screen "1牵伸相关" 1280x740, template "模板_调试"
   on GenerateScreen: "TitleUpdater"()
   IOField "IO 域_5" at 461,39 size 126x56; FormatPattern 9.999
      ProcessValue <- "ST_Cam5_Data_Var_g_tz3"
   IOField "IO 域_10" at 181,306 size 114x56; FormatPattern 9.9999
      ProcessValue <- "ST_Cam5_Data_Var_fi"
   IOField "IO 域_11" at 181,235 size 126x55; FormatPattern s9.99
      ProcessValue <- "ST_Cam5_Data_Var_g_ratioV"
   IOField "IO 域_12" at 321,235 size 126x55; FormatPattern 9.99
      ProcessValue <- "ST_Cam5_Data_Var_g_ratioT"
   TextField "文本域_13" at 181,193 size 132x43; Text 'ratioV'
   TextField "文本域_14" at 321,193 size 132x43; Text 'ratioT'
   IOField "IO 域_14" at 461,235 size 126x55; FormatPattern 9.99
      ProcessValue <- "ST_Cam5_Data_Var_g_ratio"
   TextField "文本域_16" at 461,193 size 116x43; Text 'ratio'
   IOField "IO 域_7" at 181,39 size 126x56; FormatPattern 9999
      ProcessValue <- "ST_HMI_Var_HMI_r64Position_ChuChe"
   IOField "IO 域_9" at 181,123 size 126x56; FormatPattern 9.99
      ProcessValue <- "ST_HMI_Var_HMI_r64QianShen_All"
   IOField "IO 域_13" at 321,123 size 126x56; FormatPattern 9.99
      ProcessValue <- "ST_HMI_Var_HMI_r64QianShen_First"
   IOField "IO 域_15" at 461,123 size 126x56; FormatPattern 999
      ProcessValue <- "ST_HMI_Var_HMI_r64QianShen_FirstArea"
   IOField "IO 域_16" at 601,123 size 126x56; FormatPattern 99
      ProcessValue <- "ST_HMI_Var_HMI_r64QianShen_finalArea"
   Button "Button" at 615,39 size 98x56; TextOff 'CAM5'
      Appearance <- "Cam_5_accessState"
   IOField "IO 域_8" at 321,39 size 126x56; FormatPattern 999
      ProcessValue <- "ST_Cam5_Data_Var_g_vm"
   IOField "IO 域_1" at 968,39 size 126x56; FormatPattern 9999999999
      ProcessValue <- "ST_HMI_Var_HMI_i32_ZouChe_ZhanJu_ss_1"
   IOField "IO 域_2" at 968,111 size 126x56; FormatPattern 9999
      ProcessValue <- "ST_HMI_Var_HMI_r64_ZouChe_ZhanJu_Max_20"
      Visibility <- "ST_HMI_Var_HMI_bo_ZouChe_ZhanJu_Select"
   IOField "IO 域_3" at 968,183 size 126x56; FormatPattern 9999
      ProcessValue <- "ST_HMI_Var_HMI_r64_ZouChe_ZhanJu_Max_25"
      Visibility <- "ST_HMI_Var_HMI_bo_ZouChe_ZhanJu_Select"
   IOField "IO 域_4" at 968,255 size 126x56; FormatPattern 9999
      ProcessValue <- "ST_HMI_Var_HMI_r64_ZouChe_ZhanJu_Max_30"
      Visibility <- "ST_HMI_Var_HMI_bo_ZouChe_ZhanJu_Select"
   IOField "IO 域_6" at 968,327 size 126x56; FormatPattern 9999
      ProcessValue <- "ST_HMI_Var_HMI_r64_ZouChe_ZhanJu_Max_35"
      Visibility <- "ST_HMI_Var_HMI_bo_ZouChe_ZhanJu_Select"
   IOField "IO 域_17" at 968,399 size 126x56; FormatPattern 9999
      ProcessValue <- "ST_HMI_Var_HMI_r64_ZouChe_ZhanJu_Max_40"
      Visibility <- "ST_HMI_Var_HMI_bo_ZouChe_ZhanJu_Select"
   IOField "IO 域_18" at 968,471 size 126x56; FormatPattern 9999
      ProcessValue <- "ST_HMI_Var_HMI_r64_ZouChe_ZhanJu_Max_45"
      Visibility <- "ST_HMI_Var_HMI_bo_ZouChe_ZhanJu_Select"
   IOField "IO 域_19" at 968,543 size 126x56; FormatPattern 9999
      ProcessValue <- "ST_HMI_Var_HMI_r64_ZouChe_ZhanJu_Max_Effect"
      Visibility <- "ST_HMI_Var_HMI_bo_ZouChe_ZhanJu_Select"
   Button "Button_1" at 824,111 size 126x56; TextOff '2.0米'
      on Release: SetTag("ST_HMI_Var_HMI_i16_ZouChe_ZhanJu_Select", 20)
      Visibility <- "ST_HMI_Var_HMI_bo_ZouChe_ZhanJu_Select"
      Appearance <- "ST_HMI_Var_HMI_i16_ZouChe_ZhanJu_Select"
   Button "Button_2" at 824,183 size 126x56; TextOff '2.5米'
      on Release: SetTag("ST_HMI_Var_HMI_i16_ZouChe_ZhanJu_Select", 25)
      Visibility <- "ST_HMI_Var_HMI_bo_ZouChe_ZhanJu_Select"
      Appearance <- "ST_HMI_Var_HMI_i16_ZouChe_ZhanJu_Select"
   Button "Button_3" at 824,255 size 126x56; TextOff '3.0米'
      on Release: SetTag("ST_HMI_Var_HMI_i16_ZouChe_ZhanJu_Select", 30)
      Visibility <- "ST_HMI_Var_HMI_bo_ZouChe_ZhanJu_Select"
      Appearance <- "ST_HMI_Var_HMI_i16_ZouChe_ZhanJu_Select"
   Button "Button_4" at 824,327 size 126x56; TextOff '3.5米'
      on Release: SetTag("ST_HMI_Var_HMI_i16_ZouChe_ZhanJu_Select", 35)
      Visibility <- "ST_HMI_Var_HMI_bo_ZouChe_ZhanJu_Select"
      Appearance <- "ST_HMI_Var_HMI_i16_ZouChe_ZhanJu_Select"
   Button "Button_5" at 824,399 size 126x56; TextOff '4.0米'
      on Release: SetTag("ST_HMI_Var_HMI_i16_ZouChe_ZhanJu_Select", 40)
      Visibility <- "ST_HMI_Var_HMI_bo_ZouChe_ZhanJu_Select"
      Appearance <- "ST_HMI_Var_HMI_i16_ZouChe_ZhanJu_Select"
   Button "Button_6" at 824,471 size 126x56; TextOff '4.5米'
      on Release: SetTag("ST_HMI_Var_HMI_i16_ZouChe_ZhanJu_Select", 45)
      Visibility <- "ST_HMI_Var_HMI_bo_ZouChe_ZhanJu_Select"
      Appearance <- "ST_HMI_Var_HMI_i16_ZouChe_ZhanJu_Select"
   Button "Button_7" at 824,543 size 126x56; TextOff '生效'
      Visibility <- "ST_HMI_Var_HMI_bo_ZouChe_ZhanJu_Select"
   Button "Button_8" at 181,525 size 126x56; TextOff '2.0米'; TextList "Text_list_IP_Local_Remote_Select"
      on Release: InvertBit("ST_2_HMI_bo_IP_Local_remote_Select")
      Visibility <- "ST_HMI_Var_HMI_bo_ZouChe_ZhanJu_Select"
      Appearance <- "ST_2_HMI_bo_IP_Local_remote_Select"
      ProcessValue <- "ST_2_HMI_bo_IP_Local_remote_Select"
   IOField "IO 域_21" at 327,525 size 64x56; FormatPattern 999
      ProcessValue <- "ST_2_vIPArray{0}"
      Visibility <- "ST_HMI_Var_HMI_bo_ZouChe_ZhanJu_Select"
   IOField "IO 域_22" at 398,525 size 64x56; FormatPattern 999
      ProcessValue <- "ST_2_vIPArray{1}"
      Visibility <- "ST_HMI_Var_HMI_bo_ZouChe_ZhanJu_Select"
   IOField "IO 域_23" at 470,525 size 64x56; FormatPattern 999
      ProcessValue <- "ST_2_vIPArray{2}"
      Visibility <- "ST_HMI_Var_HMI_bo_ZouChe_ZhanJu_Select"
   IOField "IO 域_24" at 542,525 size 64x56; FormatPattern 999
      ProcessValue <- "ST_2_vIPArray{3}"
      Visibility <- "ST_HMI_Var_HMI_bo_ZouChe_ZhanJu_Select"
   Button "Button_9" at 181,432 size 126x56; TextOff '设备ID'; TextList "Text_list_IP_Local_Remote_Select"
      Appearance <- "ST_2_HMI_bo_IP_Local_remote_Select"
      Visibility <- "ST_HMI_Var_HMI_bo_ZouChe_ZhanJu_Select"
      ProcessValue <- "ST_2_HMI_bo_IP_Local_remote_Select"
   IOField "IO 域_20" at 328,432 size 135x56; FormatPattern 9999
      ProcessValue <- "ST_HMI_Var_HMI_u32_DeviceID"
      Visibility <- "ST_HMI_Var_HMI_bo_ZouChe_ZhanJu_Select"

screen "2加捻相关" 1280x740, template "模板_调试"
   on GenerateScreen: "TitleUpdater"()
   TextField "Text Field_58" at 327,45 size 304x42; Text '锭子加捻加速度'
   TextField "Text Field_1" at 168,8 size 156x23; Text '一、锭子加捻TO参数:'
   TextField "Text Field_60" at 327,101 size 304x42; Text '锭子加捻正起始加加速度'
   TextField "Text Field_61" at 327,157 size 304x42; Text '锭子加捻正终止加加速度'
   TextField "Text Field_62" at 327,213 size 304x42; Text '锭子加捻负起始加加速度'
   TextField "Text Field_63" at 327,269 size 304x42; Text '锭子加捻负终止加加速度'
   TextField "Text Field_66" at 327,325 size 304x42; Text '锭子点动加捻加速度'
   IOField "IO Field_38" at 194,41 size 112x42; FormatPattern 99999
      ProcessValue <- "ST_HMI_Var_HMI_r64Axis_DingZi_PositiveAccel_JiaNian"
   IOField "IO Field_40" at 194,97 size 112x42; FormatPattern 99999
      ProcessValue <- "ST_HMI_Var_HMI_r64Axis_DingZi_Positiveaccelstartjerk_JiaNian"
   IOField "IO Field_41" at 194,153 size 112x42; FormatPattern 99999
      ProcessValue <- "ST_HMI_Var_HMI_r64Axis_DingZi_positiveaccelendjerk_JiaNian"
   IOField "IO Field_42" at 194,209 size 112x42; FormatPattern 99999
      ProcessValue <- "ST_HMI_Var_HMI_r64Axis_DingZi_negativeaccelstartjerk_JiaNian"
   IOField "IO Field_43" at 194,265 size 112x42; FormatPattern 99999
      ProcessValue <- "ST_HMI_Var_HMI_r64Axis_DingZi_negativeaccelendjerk_JiaNian"
   IOField "IO Field_44" at 194,321 size 112x42; FormatPattern 99999
      ProcessValue <- "ST_HMI_Var_HMI_r64AccVelocity_Jog_JiaNian"

screen "3退绕相关1" 1280x740, template "模板_调试"
   on GenerateScreen: "TitleUpdater"()
   TextField "Text Field_58" at 153,27 size 668x41; Text '1.退绕成形弓速度————————————'
   TextField "Text Field_59" at 153,77 size 668x41; Text '2.退绕成形弓加速度————————————'
   TextField "Text Field_60" at 153,128 size 668x40; Text '3.退绕成形弓正向开始加加速度————————————'
   TextField "Text Field_61" at 153,178 size 668x41; Text '4.退绕成形弓正向结束加加速度————————————'
   TextField "Text Field_62" at 153,229 size 668x40; Text '5.退绕成形弓反向开始加加速度————————————'
   TextField "Text Field_1" at 153,5 size 247x26; Text '一、退绕成形弓TO参数:'
   TextField "Text Field_63" at 153,279 size 668x41; Text '6.退绕成形弓反向结束加加速度————————————'
   TextField "Text Field_41" at 153,361 size 668x41; Text '1.退绕结束纱线提前角度（越大，卷绕时，包络层螺距越大）—————————————————————'
   TextField "Text Field_42" at 153,413 size 668x41; Text '2.退绕开始位置—————————————————————————————'
   TextField "Text Field_43" at 153,465 size 668x41; Text '3.退绕结束位置—————————————————————————'
   TextField "Text Field_44" at 153,517 size 668x41; Text '4.退绕拐点比例———————————————————————————'
   TextField "Text Field_45" at 153,569 size 668x41; Text '5.退绕拐点点数---------------------'
   TextField "Text Field_3" at 153,327 size 260x26; Text '二、Cam_3曲线计算参数:'
   TextField "Text Field_46" at 153,621 size 668x41; Text '6.退绕圈数比例（越大，圈数越多，一般以0.03为单位调整）---------------------'
   IOField "IO Field_39" at 819,23 size 109x41; FormatPattern 9999
      ProcessValue <- "ST_HMI_Var_HMI_r64Axis_ChengXing_Velocity_TuiRao"
   IOField "IO Field_43" at 819,74 size 109x41; FormatPattern 9999
      ProcessValue <- "ST_HMI_Var_HMI_r64Axis_ChengXing_PositiveAccel_TuiRao"
   IOField "IO Field_44" at 819,125 size 109x41; FormatPattern 9999
      ProcessValue <- "ST_HMI_Var_HMI_r64Axis_ChengXing_positiveaccelstartjerk_TuiRao"
   IOField "IO Field_45" at 819,177 size 109x41; FormatPattern 9999
      ProcessValue <- "ST_HMI_Var_HMI_r64Axis_ChengXing_positiveaccelendjerk_TuiRao"
   IOField "IO Field_46" at 819,228 size 109x41; FormatPattern 9999
      ProcessValue <- "ST_HMI_Var_HMI_r64Axis_ChengXing_negativeaccelstartjerk_TuiRao"
   IOField "IO Field_47" at 819,280 size 109x40; FormatPattern 9999
      ProcessValue <- "ST_HMI_Var_HMI_r64Axis_ChengXing_negativeaccelendjerk_TuiRao"
   IOField "IO Field_53" at 819,367 size 109x41; FormatPattern 9999
      ProcessValue <- "ST_HMI_Var_HMI_alpha_TuiRao_5"
   IOField "IO Field_54" at 819,468 size 109x41; FormatPattern 99999
      ProcessValue <- "ST_HMI_Var_HMI_x_TuiRao_5"
   IOField "IO Field_55" at 819,570 size 109x41; FormatPattern 99
      ProcessValue <- "ST_HMI_Var_HMI_n_Change_TuiRao"
   IOField "IO Field_56" at 819,417 size 109x41; FormatPattern 9999
      ProcessValue <- "ST_HMI_Var_HMI_x_TuiRao_0"
   IOField "IO Field_57" at 819,519 size 109x41; FormatPattern 9.99
      ProcessValue <- "ST_HMI_Var_HMI_k_TuiRao"
   IOField "IO Field_58" at 819,621 size 109x41; FormatPattern 9.99
      ProcessValue <- "ST_HMI_Var_HMI_scalevalue_Cam_3"

screen "4退绕相关2" 1280x740, template "模板_调试"
   on GenerateScreen: "TitleUpdater"()
   TextField "Text Field_48" at 151,98 size 786x42; Text '2.退绕锭子响应正向加速度————————————————————'
   TextField "Text Field_49" at 151,154 size 786x42; Text '3.退绕锭子响应反向加速度————————————————————————'
   TextField "Text Field_1" at 151,9 size 204x27; Text '三、cam_3 TO参数'
   TextField "Text Field_65" at 151,42 size 786x42; Text '1.退绕锭子响应速度————————————————————'
   TextField "Text Field_4" at 151,210 size 235x27; Text '四、退绕张力TO参数'
   TextField "Text Field_54" at 151,309 size 786x42; Text '2.退绕张力加速度比例————————————————————'
   TextField "Text Field_66" at 151,253 size 786x42; Text '1.退绕张力速度比例————————————————————'
   TextField "Text Field_5" at 151,407 size 377x27; Text '五、退绕工艺进程衔接紧密性参数:'
   TextField "Text Field_63" at 151,449 size 786x42; Text '1.退绕锭子速度减少值————————————————————'
   TextField "Text Field_64" at 151,505 size 786x42; Text '2.开始退绕锭子速度————————————'
   IOField "IO Field_40" at 935,42 size 112x42; FormatPattern 9999
      ProcessValue <- "ST_HMI_Var_HMI_r64_cam_DingZi_velocity_TuiRao"
   IOField "IO Field_43" at 935,98 size 112x42; FormatPattern 99999
      ProcessValue <- "ST_HMI_Var_HMI_r64_cam_DingZi_positiveaccel_TuiRao"
   IOField "IO Field_47" at 935,154 size 112x42; FormatPattern 99999
      ProcessValue <- "ST_HMI_Var_HMI_r64_cam_DingZi_negativeaccel_TuiRao"
   IOField "IO Field_50" at 935,253 size 112x42; FormatPattern 9.99
      ProcessValue <- "ST_HMI_Var_HMI_r64Axis_1_ZhangLi_Velocity_from_ChengXing_ratio_tuirao"
   IOField "IO Field_51" at 935,309 size 112x42; FormatPattern 9.99
      ProcessValue <- "ST_HMI_Var_HMI_r64Axis_1_ZhangLi_PositiveAccel_from_ChengXing_ratio_tuirao"
   IOField "IO Field_52" at 935,449 size 112x42; FormatPattern 9999
      ProcessValue <- "ST_HMI_Var_HMI_r64Axis_DingZi_Velocity_JianShaoZhi"
   IOField "IO Field_53" at 935,505 size 112x42; FormatPattern 99
      ProcessValue <- "ST_HMI_Var_HMI_r64Axis_DingZi_Velocity_Start_TuiRao"
   IOField "IO Field_56" at 935,365 size 112x42; FormatPattern 9.99
      ProcessValue <- "ST_HMI_Var_HMI_r64Axis_1_ZhangLi_Additive_Torque_TuiRao"

screen "5成形相关" 1280x740, template "模板_调试"
   on GenerateScreen: "TitleUpdater"()
   TextField "Text Field_1" at 140,1 size 267x29; Text '一、成形凸轮曲线计算参数:'
   TextField "Text Field_58" at 138,36 size 648x39; Text '1.卷绕提前角度1——————————————————————'
   TextField "Text Field_59" at 138,81 size 648x40; Text '2.卷绕提前角度2——————————————————————————'
   TextField "Text Field_60" at 138,127 size 648x40; Text '3.卷绕提前角度3——————————————————————————'
   TextField "Text Field_61" at 138,174 size 648x40; Text '4.生头开始上锥体高度修正值——————————————————————————'
   TextField "Text Field_62" at 138,220 size 648x39; Text '5.最大直径时上椎体高度修正值——————————————————————————'
   TextField "Text Field_63" at 139,266 size 648x39; Text '6.满纱时上椎体高度修正值————————————————————————'
   TextField "Text Field_2" at 140,308 size 165x29; Text '二、cam1TO参数:'
   TextField "Text Field_64" at 140,337 size 648x39; Text '1.卷绕成形响应速度——————————————————————'
   TextField "Text Field_65" at 140,385 size 648x40; Text '2.卷绕成形响应正向加速度——————————————————————————'
   TextField "Text Field_66" at 140,435 size 648x40; Text '3.卷绕成形响应负向加速度——————————————————————————'
   TextField "Text Field_67" at 140,485 size 648x40; Text '4.卷绕成形响应正向开始加加速度——————————————————————————'
   TextField "Text Field_68" at 140,535 size 648x39; Text '5.卷绕成形响应正向结束加加速度——————————————————————————'
   TextField "Text Field_69" at 140,584 size 649x39; Text '6.卷绕成形响应反向开始加加速度————————————————————————'
   TextField "Text Field_70" at 140,633 size 648x40; Text '7.卷绕成形响应反向结束加加速度————————————————————————'
   IOField "IO Field_51" at 786,32 size 106x40; FormatPattern 99.9
      ProcessValue <- "ST_HMI_Var_HMI_alpha_JuanRao_1"
   IOField "IO Field_52" at 786,337 size 106x39; FormatPattern 9999
      ProcessValue <- "ST_HMI_Var_HMI_r64_cam_ChengXing_velocity_juanrao"
   IOField "IO Field_53" at 786,79 size 106x40; FormatPattern 99.9
      ProcessValue <- "ST_HMI_Var_HMI_alpha_JuanRao_2"
   IOField "IO Field_54" at 786,126 size 106x40; FormatPattern 99.9
      ProcessValue <- "ST_HMI_Var_HMI_alpha_JuanRao_3"
   IOField "IO Field_55" at 786,173 size 106x39; FormatPattern 99.9
      ProcessValue <- "ST_HMI_Var_HMI_r64_Hs2_0_delt"
   IOField "IO Field_56" at 786,219 size 106x39; FormatPattern 99.9
      ProcessValue <- "ST_HMI_Var_HMI_r64_Hs2_D_delt"
   IOField "IO Field_57" at 786,266 size 106x40; FormatPattern 99.9
      ProcessValue <- "ST_HMI_Var_HMI_r64_Hs2_N_delt"
   IOField "IO Field_58" at 786,385 size 106x40; FormatPattern 9999
      ProcessValue <- "ST_HMI_Var_HMI_r64_cam_ChengXing_positiveaccel_juanrao"
   IOField "IO Field_59" at 786,435 size 106x40; FormatPattern 9999
      ProcessValue <- "ST_HMI_Var_HMI_r64_cam_ChengXing_negativeaccel_juanrao"
   IOField "IO Field_60" at 786,485 size 106x40; FormatPattern 9999
      ProcessValue <- "ST_HMI_Var_HMI_r64_cam_ChengXing_positiveaccelstartjerk_juanrao"
   IOField "IO Field_61" at 786,535 size 106x39; FormatPattern 9999
      ProcessValue <- "ST_HMI_Var_HMI_r64_cam_ChengXing_positiveaccelendjerk_juanrao"
   IOField "IO Field_62" at 786,584 size 106x39; FormatPattern 9999
      ProcessValue <- "ST_HMI_Var_HMI_r64_cam_ChengXing_negativeaccelstartjerk_juanrao"
   IOField "IO Field_63" at 786,633 size 106x40; FormatPattern 9999
      ProcessValue <- "ST_HMI_Var_HMI_r64_cam_ChengXing_negativeaccelendjerk_juanrao"

screen "6卷绕相关1" 1280x740, template "模板_调试"
   on GenerateScreen: "TitleUpdater"()
   TextField "Text Field_1" at 155,9 size 224x32; Text '一、锭子卷绕TO参数:'
   TextField "Text Field_58" at 155,42 size 786x42; Text '1.卷绕锭子最小速度————————————————————————'
   TextField "Text Field_63" at 155,98 size 786x42; Text '2.卷绕锭子最大速度————————————————————————'
   TextField "Text Field_64" at 155,154 size 786x42; Text '3.卷绕锭子加速度————————————————————————'
   TextField "Text Field_2" at 155,210 size 224x32; Text '二、卷绕张力TO参数:'
   TextField "Text Field_59" at 155,252 size 786x42; Text '1.卷绕张力速度————————————————————————'
   TextField "Text Field_67" at 155,308 size 786x42; Text '2.卷绕张力附加力矩————————————————————————'
   IOField "IO Field_38" at 939,42 size 112x42; FormatPattern 999
      ProcessValue <- "ST_HMI_Var_HMI_r64Axis_DingZi_Velocity_JuanRao_min"
   IOField "IO Field_41" at 939,98 size 112x42; FormatPattern 99999
      ProcessValue <- "ST_HMI_Var_HMI_r64Axis_DingZi_Velocity_JuanRao_max"
   IOField "IO Field_46" at 939,154 size 112x42; FormatPattern 99999
      ProcessValue <- "ST_HMI_Var_HMI_r64Axis_DingZi_PositiveAccel_JuanRao"
   IOField "IO Field_39" at 939,252 size 112x42; FormatPattern 99.9
      ProcessValue <- "ST_HMI_Var_HMI_r64Axis_1_ZhangLi_Velocity_JuanRao"
   IOField "IO Field_40" at 939,308 size 112x42; FormatPattern 9.99
      ProcessValue <- "ST_HMI_Var_HMI_r64Axis_1_ZhangLi_Additive_Torque_JuanRao"

screen "7卷绕相关2" 1280x740, template "模板_调试"
   on GenerateScreen: "TitleUpdater"()
   TextField "Text Field_37" at 221,161 size 286x41; Text '刚生头时卷绕中间调整值————————————'
   TextField "Text Field_38" at 221,215 size 286x41; Text '刚生头时卷绕到底调整值————————————'
   TextField "Text Field_39" at 221,107 size 286x41; Text '满纱时张力弓位置————————————'
   TextField "Text Field_40" at 221,53 size 286x41; Text '最大直径时张力弓位置————————————'
   TextField "Text Field_41" at 221,0 size 286x41; Text '刚生头时张力弓位置————————————'
   TextField "Text Field_42" at 221,269 size 286x41; Text '卷绕张力弓中间位置修正————————————'
   TextField "Text Field_43" at 221,323 size 286x41; Text '卷绕张力弓到底位置修正------------'
   TextField "Text Field_44" at 221,377 size 286x41; Text '卷绕张力弓开始位置修正————————————'
   TextField "Text Field_45" at 221,431 size 286x41; Text '张力弓反馈系数————————————'
   TextField "Text Field_47" at 221,538 size 286x41; Text '卷绕锭子设定走车位置——————————————————'
   TextField "Text Field_51" at 642,0 size 286x41; Text '中间调整最小值————————————'
   TextField "Text Field_52" at 642,54 size 286x41; Text '中间调整最小增量值————————————'
   TextField "Text Field_53" at 642,108 size 286x41; Text '中间调整最大增量值————————————'
   TextField "Text Field_54" at 642,161 size 286x41; Text '中间调整系数————————————'
   TextField "Text Field_55" at 642,215 size 286x41; Text '到底调整最小值————————————'
   TextField "Text Field_56" at 642,269 size 286x41; Text '到底调整最小增量值————————————'
   TextField "Text Field_57" at 642,323 size 286x41; Text '到底调整最大增量值————————————'
   TextField "Text Field_59" at 642,377 size 286x41; Text '到底调整系数————————————'
   TextField "Text Field_60" at 642,431 size 286x41; Text '张力中央采样位置————————————'
   IOField "IO Field_20" at 507,161 size 108x41; FormatPattern 99.99
      ProcessValue <- "ST_HMI_Var_HMI_f1_n_delt_new_0"
   IOField "IO Field_21" at 507,215 size 108x41; FormatPattern 99.99
      ProcessValue <- "ST_HMI_Var_HMI_g1_n_delt_new_0"
   IOField "IO Field_22" at 507,108 size 108x40; FormatPattern 99.99
      ProcessValue <- "ST_HMI_Var_HMI_r64Axis_1_ZhangLi_Position_JuanRao_Set_N"
   IOField "IO Field_23" at 507,54 size 108x40; FormatPattern 99.99
      ProcessValue <- "ST_HMI_Var_HMI_r64Axis_1_ZhangLi_Position_JuanRao_Set_ND"
   IOField "IO Field_24" at 507,0 size 108x40; FormatPattern 99.99
      ProcessValue <- "ST_HMI_Var_HMI_r64Axis_1_ZhangLi_Position_JuanRao_Set_0"
   IOField "IO Field_25" at 507,269 size 108x40; FormatPattern 99.99
      ProcessValue <- "ST_HMI_Var_HMI_f1_n_ZhangLi_Set_PianTiao_0"
   IOField "IO Field_26" at 507,323 size 108x40; FormatPattern 99.99
      ProcessValue <- "ST_HMI_Var_HMI_g1_n_ZhangLi_Set_PianTiao_0"
   IOField "IO Field_27" at 507,377 size 108x40; FormatPattern 99.99
      ProcessValue <- "ST_HMI_Var_HMI_gam_ZhangLi_Set_PianTiao_0"
   IOField "IO Field_28" at 507,431 size 108x40; FormatPattern 99.99
      ProcessValue <- "ST_HMI_Var_HMI_r64_k_ZhangLi_Rate"
   IOField "IO Field_30" at 507,538 size 108x41; FormatPattern 99.99
      ProcessValue <- "ST_VAR_ZouChe_g_r64Axis_ZouChe_Position_JuanRao_DingZi_Velocity_Set"
   IOField "IO Field_34" at 928,0 size 108x40; FormatPattern 99.99
      ProcessValue <- "ST_FC_Var_g_f1_n_piantiao_min"
   IOField "IO Field_35" at 928,54 size 108x40; FormatPattern 99.99
      ProcessValue <- "ST_FC_Var_g_f1_n_delt_min"
   IOField "IO Field_36" at 928,108 size 108x40; FormatPattern 99.99
      ProcessValue <- "ST_FC_Var_g_f1_n_delt_max"
   IOField "IO Field_37" at 928,161 size 108x41; FormatPattern 99.99
      ProcessValue <- "ST_FC_Var_g_f1_n_delt_ratio"
   IOField "IO Field_38" at 928,215 size 108x41; FormatPattern 99.99
      ProcessValue <- "ST_FC_Var_g_g1_n_piantiao_min"
   IOField "IO Field_39" at 928,269 size 108x40; FormatPattern 99.99
      ProcessValue <- "ST_FC_Var_g_g1_n_delt_min"
   IOField "IO Field_40" at 928,323 size 108x40; FormatPattern 99.99
      ProcessValue <- "ST_FC_Var_g_g1_n_delt_max"
   IOField "IO Field_42" at 928,377 size 108x40; FormatPattern 99.99
      ProcessValue <- "ST_FC_Var_g_g1_n_delt_ratio"
   IOField "IO Field_43" at 928,431 size 108x40; FormatPattern 9999
      ProcessValue <- "ST_FC_Var_g_Position_ZouChe_Zhangli_mid"

screen "8存绕相关" 1280x740, template "模板_调试"
   on GenerateScreen: "TitleUpdater"()
   TextField "Text Field_41" at 152,454 size 430x40; Text '存绕锭子加速度------------'
   TextField "Text Field_42" at 152,508 size 430x40; Text '存绕锭子加速度比例————————————'
   TextField "Text Field_43" at 152,10 size 430x40; Text '存绕成形速度------------'
   TextField "Text Field_44" at 152,64 size 430x40; Text '存绕成形加速度————————————'
   TextField "Text Field_45" at 152,118 size 430x40; Text '存绕成形正向开始加加速度————————————'
   TextField "Text Field_48" at 152,171 size 430x41; Text '存绕成形正向结束加加速度————————————'
   TextField "Text Field_49" at 152,225 size 430x41; Text '存绕成形反向开始加加速度————————————'
   TextField "Text Field_50" at 152,279 size 430x40; Text '存绕成形反向结束加加速度————————————'
   TextField "Text Field_51" at 152,333 size 430x40; Text '存绕长度————————————————'
   TextField "Text Field_52" at 152,387 size 430x40; Text '存绕走车增量————————————————'
   IOField "IO Field_24" at 582,454 size 108x40; FormatPattern 99999
      ProcessValue <- "ST_Main_Var_g_r64Axis_DingZi_PositiveAccel_CunRao"
   IOField "IO Field_25" at 582,508 size 108x40; FormatPattern 99.99
      ProcessValue <- "ST_Main_Var_g_r64Axis_DingZi_Velocity_CunRao_ratio"
   IOField "IO Field_26" at 582,10 size 108x40; FormatPattern 999
      ProcessValue <- "ST_HMI_Var_HMI_r64Axis_ChengXing_Velocity_CunRao"
   IOField "IO Field_27" at 582,64 size 108x40; FormatPattern 9999
      ProcessValue <- "ST_HMI_Var_HMI_r64Axis_ChengXing_PositiveAccel_CunRao"
   IOField "IO Field_28" at 582,118 size 108x40; FormatPattern 99999
      ProcessValue <- "ST_HMI_Var_HMI_r64Axis_ChengXing_positiveaccelstartjerk_CunRao"
   IOField "IO Field_31" at 582,171 size 108x41; FormatPattern 99999
      ProcessValue <- "ST_HMI_Var_HMI_r64Axis_ChengXing_positiveaccelendjerk_CunRao"
   IOField "IO Field_32" at 582,225 size 108x41; FormatPattern 99999
      ProcessValue <- "ST_HMI_Var_HMI_r64Axis_ChengXing_negativeaccelstartjerk_CunRao"
   IOField "IO Field_33" at 582,279 size 108x40; FormatPattern 99999
      ProcessValue <- "ST_HMI_Var_HMI_r64Axis_ChengXing_negativeaccelendjerk_CunRao"
   IOField "IO Field_34" at 582,333 size 108x40; FormatPattern 99
      ProcessValue <- "ST_HMI_Var_HMI_r64_Lcr"
   IOField "IO Field_35" at 582,387 size 108x40; FormatPattern 99
      ProcessValue <- "ST_HMI_Var_HMI_r64_Delt_Position_ZouChe_Cam_1_CunRao"

screen "9自动停止" 1280x740, template "模板_调试"
   on GenerateScreen: "TitleUpdater"()
   TextField "Text Field_1" at 159,6 size 178x32; Text '一、走车TO参数:'
   TextField "Text Field_58" at 159,43 size 688x42; Text '1.自动停止走车位置————————————————————————'
   TextField "Text Field_59" at 159,99 size 688x42; Text '2.自动停止走车速度————————————————————————'
   TextField "Text Field_60" at 159,155 size 688x42; Text '3.自动停止走车加速度————————————————————————'
   TextField "Text Field_61" at 159,253 size 688x42; Text '1.自动停止锭子加速度————————————————————————'
   TextField "Text Field_62" at 159,350 size 688x42; Text '1.自动停止总牵伸————————————————————————'
   TextField "Text Field_63" at 159,407 size 688x42; Text '2.自动停止无捻牵伸————————————————————————'
   TextField "Text Field_64" at 159,463 size 688x42; Text '3.自动停止分散牵伸————————————————————————'
   TextField "Text Field_65" at 159,519 size 688x42; Text '4.自动停止设定捻度————————————————————————'
   TextField "Text Field_2" at 159,207 size 178x32; Text '二、锭子TO参数:'
   TextField "Text Field_3" at 159,305 size 200x32; Text '三、工艺参数设置:'
   TextField "Text Field_66" at 159,575 size 688x42; Text '5.自动停止设定捻速————————————————————————'
   IOField "IO Field_38" at 845,39 size 112x42; FormatPattern 99999
      ProcessValue <- "ST_HMI_Var_HMI_r64Axis_ZouChe_Position_ZiDongTingZhi"
   IOField "IO Field_39" at 845,95 size 112x42; FormatPattern 99999
      ProcessValue <- "ST_HMI_Var_HMI_r64Axis_ZouChe_Velocity_ZiDongTingZhi"
   IOField "IO Field_40" at 845,151 size 112x42; FormatPattern 99999
      ProcessValue <- "ST_HMI_Var_HMI_r64Axis_ZouChe_PositiveAccel_ZiDongTingZhi"
   IOField "IO Field_41" at 845,249 size 112x42; FormatPattern 99999
      ProcessValue <- "ST_HMI_Var_HMI_r64Axis_DingZi_PositiveAccel_ZiDongTingZhi"
   IOField "IO Field_42" at 845,347 size 112x42; FormatPattern 9.999
      ProcessValue <- "ST_HMI_Var_HMI_r64_ZiDongTingZhi_QianShen_All"
   IOField "IO Field_43" at 845,403 size 112x42; FormatPattern 9.999
      ProcessValue <- "ST_HMI_Var_HMI_r64_ZiDongTingZhi_QianShen_WuNian"
   IOField "IO Field_44" at 845,459 size 112x42; FormatPattern 9.999
      ProcessValue <- "ST_HMI_Var_HMI_r64_ZiDongTingZhi_QianShen_FenSan"
   IOField "IO Field_45" at 845,515 size 112x42; FormatPattern 99999
      ProcessValue <- "ST_HMI_Var_HMI_r64_ZiDongTingZhi_NianDu_SheDing"
   IOField "IO Field_46" at 845,571 size 112x42; FormatPattern 99999
      ProcessValue <- "ST_HMI_Var_HMI_r64_ZiDongTingZhi_NianSu_SheDing"

screen "10走车相关" 1280x740, template "模板_调试"
   on GenerateScreen: "TitleUpdater"()
   TextField "Text Field_37" at 390,93 size 242x40; Text '出车正加速度'
   TextField "Text Field_38" at 390,228 size 242x40; Text '出车正起始加加速度'
   TextField "Text Field_39" at 851,93 size 227x40; Text '进车加速度'
   TextField "Text Field_40" at 390,297 size 242x40; Text '出车正终止加加速度'
   TextField "Text Field_41" at 390,364 size 242x42; Text '出车负起始加加速度'
   TextField "Text Field_42" at 390,433 size 242x40; Text '出车负终止加加速度'
   TextField "Text Field_43" at 851,367 size 227x40; Text '进车负终止加加速度'
   TextField "Text Field_44" at 851,298 size 227x42; Text '进车负起始加加速度'
   TextField "Text Field_45" at 851,231 size 227x40; Text '进车正终止加加速度'
   TextField "Text Field_46" at 851,162 size 227x40; Text '进车正起始加加速度'
   TextField "Text Field_47" at 390,24 size 242x42; Text '出车速度'
   TextField "Text Field_48" at 851,24 size 227x42; Text '进车速度'
   IOField "IO Field_56" at 245,93 size 114x40; FormatPattern 9999
      ProcessValue <- "ST_HMI_Var_HMI_r64PositiveAccel_ZouChe_ChuChe"
   IOField "IO Field_69" at 244,228 size 114x40; FormatPattern 9999999
      ProcessValue <- "ST_HMI_Var_HMI_r64Axis_ZouChe_positiveaccelstartjerk_ChuChe"
   IOField "IO Field_70" at 699,93 size 108x40; FormatPattern 9999
      ProcessValue <- "ST_HMI_Var_HMI_r64PositiveAccel_ZouChe_JinChe"
   IOField "IO Field_75" at 243,297 size 114x40; FormatPattern 9999999
      ProcessValue <- "ST_HMI_Var_HMI_r64Axis_ZouChe_positiveaccelendjerk_ChuChe"
   IOField "IO Field_78" at 244,364 size 114x42; FormatPattern 9999999
      ProcessValue <- "ST_HMI_Var_HMI_r64Axis_ZouChe_negativeaccelstartjerk_ChuChe"
   IOField "IO Field_79" at 244,433 size 114x40; FormatPattern 9999999
      ProcessValue <- "ST_HMI_Var_HMI_r64Axis_ZouChe_negativeaccelendjerk_ChuChe"
   IOField "IO Field_80" at 699,231 size 108x40; FormatPattern 9999999
      ProcessValue <- "ST_HMI_Var_HMI_r64Axis_ZouChe_positiveaccelendjerk_JinChe"
   IOField "IO Field_81" at 699,298 size 108x42; FormatPattern 9999999
      ProcessValue <- "ST_HMI_Var_HMI_r64Axis_ZouChe_negativeaccelstartjerk_JinChe"
   IOField "IO Field_82" at 699,367 size 108x40; FormatPattern 9999999
      ProcessValue <- "ST_HMI_Var_HMI_r64Axis_ZouChe_negativeaccelendjerk_JinChe"
   IOField "IO Field_83" at 699,162 size 108x40; FormatPattern 9999999
      ProcessValue <- "ST_HMI_Var_HMI_r64Axis_ZouChe_positiveaccelstartjerk_JinChe"
   IOField "IO Field_57" at 245,24 size 114x42; FormatPattern 9999
      ProcessValue <- "ST_HMI_Var_HMI_r64Velocity_ChuChe"
   IOField "IO Field_84" at 699,24 size 108x42; FormatPattern 9999
      ProcessValue <- "ST_HMI_Var_HMI_r64Velocity_JinChe"
   TextField "Text Field_1" at 390,159 size 242x40; Text '出车负加速度'
   IOField "IO Field_1" at 245,159 size 114x40; FormatPattern 9999
      ProcessValue <- "ST_HMI_Var_HMI_r64NegativeAccel_ZouChe_ChuChe"

screen "11生头相关" 1280x740, template "模板_调试"
   on GenerateScreen: "TitleUpdater"()
   IOField "IO Field_41" at 266,24 size 112x42; FormatPattern 99
      ProcessValue <- "ST_HMI_Var_HMI_r64_MaoZhou_TouShu"
   IOField "IO Field_46" at 266,432 size 112x42; FormatPattern 999
      ProcessValue <- "ST_HMI_Var_HMI_r64Axis_ZouChe_Position_KongDing_8"
   IOField "IO Field_1" at 266,80 size 112x42; FormatPattern 99
      ProcessValue <- "ST_HMI_Var_HMI_r64Axis_ChengXing_Position_delt_KongDing_8"
   IOField "IO Field_2" at 266,544 size 112x42; FormatPattern 99.9
      ProcessValue <- "ST_HMI_Var_HMI_r64_DingZi_Zouche_ratio_KongDing_9"
   IOField "IO Field_3" at 522,432 size 112x42; FormatPattern 999
      ProcessValue <- "ST_HMI_Var_HMI_r64Axis_ZouChe_Position_LuoSha_8"
   IOField "IO Field_4" at 522,544 size 112x42; FormatPattern 99.9
      ProcessValue <- "ST_HMI_Var_HMI_r64_DingZi_Zouche_ratio_LuoSha_9"
   IOField "IO Field_6" at 266,488 size 112x42; FormatPattern 999
      ProcessValue <- "ST_HMI_Var_HMI_r64Axis_ZouChe_Position_KongDing_9"
   IOField "IO Field_5" at 458,488 size 112x42; FormatPattern 999
      ProcessValue <- "ST_HMI_Var_HMI_r64Axis_ZouChe_Position_LuoSha_9"
   IOField "IO Field_7" at 266,136 size 112x42; FormatPattern 999.9
      ProcessValue <- "ST_HMI_Var_HMI_r64Position_ChuChe_KongDing_65"
   IOField "IO Field_8" at 266,192 size 112x42; FormatPattern 9.99
      ProcessValue <- "ST_HMI_Var_HMI_r64QianShen_KongDing_65"
   IOField "IO Field_9" at 266,248 size 112x42; FormatPattern 99.9
      ProcessValue <- "ST_HMI_Var_HMI_r64_DingZi_Zouche_ratio_KongDing_65"
   IOField "IO Field_10" at 266,304 size 112x42; FormatPattern 99.9
      ProcessValue <- "ST_HMI_Var_HMI_r64Axis_ZouChe_Position_ShengTou_Start_Position"
   IOField "IO Field_11" at 394,432 size 112x42; FormatPattern 999
      ProcessValue <- "ST_HMI_Var_HMI_r64Axis_ZouChe_Position_KongDing_8_1"
   IOField "IO Field_12" at 394,544 size 112x42; FormatPattern 99.9
      ProcessValue <- "ST_HMI_Var_HMI_r64_DingZi_Zouche_ratio_KongDing_9_1"
   TextField "Text Field_8" at 404,24 size 332x42; Text '1.毛轴头数'
   TextField "Text Field_9" at 404,80 size 332x42; Text '2.成形弓上升量'
   TextField "Text Field_10" at 650,432 size 264x42; Text '7.走车第一次回车量'
   TextField "Text Field_11" at 650,488 size 264x42; Text '8.纱管底部纱线卷绕长度'
   TextField "Text Field_12" at 650,544 size 264x42; Text '9.锭子走车传动比'
   TextField "Text Field_16" at 404,136 size 332x42; Text '3.回绕出车展距'
   TextField "Text Field_17" at 404,192 size 332x42; Text '4.回绕牵伸'
   TextField "Text Field_18" at 404,248 size 332x42; Text '5.回绕锭子走车传动比'
   TextField "Text Field_1" at 404,304 size 332x42; Text '6.生头起点位置'
   TextField "Text Field_2" at 266,392 size 112x32; Text '空锭(先插管)'
   TextField "Text Field_3" at 394,392 size 112x32; Text '空锭(光锭)'
   TextField "Text Field_4" at 522,392 size 112x32; Text '落纱生头'
   Button "OBJECT_6" at 892,161 size 170x66; TextOff '拔锭脚纱选择 / EXIT'
      on Release: InvertBit("ST_HMI_Var_HMI_bo_BaShaTou_Select")
      Visibility <- "ST_HMI_Var_HMI_i16_ShengTou_Select"
      Appearance <- "ST_HMI_Var_HMI_bo_BaShaTou_Select"
      ObjectEnable <- "ST_Main_Var_g_i16_KongDing_Status"
   IOField "IO Field_13" at 893,116 size 168x42; Authorization "User administration"; FormatPattern 99
      ProcessValue <- "ST_HMI_Var_HMI_r64Axis_ZouChe_Position_LuoSha_112_Delta_BaTou"
      Visibility <- "ST_HMI_Var_HMI_i16_ShengTou_Select"
   TextField "Text Field_5" at 892,77 size 170x38; Text '补偿距离'
      Visibility <- "ST_HMI_Var_HMI_i16_ShengTou_Select"

screen "12张力弓整定" 1280x740, template "模板_调试"
   on GenerateScreen: "TitleUpdater"()
   Button "OBJECT_109" at 249,47 size 182x70; TextOff '张力测定 / EXIT'
      on Press: SetTag("ST_Main_Var_g_i16_Mode_Selected", 256)
      Appearance <- "ST_Main_Var_g_bo_Mode_Enabled_Manual"
   Button "OBJECT_110" at 249,233 size 182x70; TextOff '张力测定启动 / EXIT'
      on Release: ResetBit("ST_HMI_Var_HMI_bo_ZhangLi_CeDing_Start")
      on Press: SetBit("ST_HMI_Var_HMI_bo_ZhangLi_CeDing_Start")
      Appearance <- "ST_Main_Var_g_bo_Mode_Enabled_Manual"
   IOField "I/O 域_1" at 631,41 size 86x40; FormatPattern 99.99
      ProcessValue <- "ST_Var_ZLCD_HMI_r64Axis_1_ZhangLi_Torque_CeDing_N{0}"
   IOField "I/O 域_2" at 631,85 size 86x40; FormatPattern 99.99
      ProcessValue <- "ST_Var_ZLCD_HMI_r64Axis_1_ZhangLi_Torque_CeDing_N{1}"
   IOField "I/O 域_3" at 631,129 size 86x40; FormatPattern 99.99
      ProcessValue <- "ST_Var_ZLCD_HMI_r64Axis_1_ZhangLi_Torque_CeDing_N{2}"
   IOField "I/O 域_4" at 631,173 size 86x40; FormatPattern 99.99
      ProcessValue <- "ST_Var_ZLCD_HMI_r64Axis_1_ZhangLi_Torque_CeDing_N{3}"
   IOField "I/O 域_5" at 631,217 size 86x40; FormatPattern 99.99
      ProcessValue <- "ST_Var_ZLCD_HMI_r64Axis_1_ZhangLi_Torque_CeDing_N{4}"
   IOField "I/O 域_6" at 631,260 size 86x40; FormatPattern 99.99
      ProcessValue <- "ST_Var_ZLCD_HMI_r64Axis_1_ZhangLi_Torque_CeDing_N{6}"
   Button "按钮_1" at 855,256 size 136x44; TextOff '调整'
      on Release: ResetBit("ST_Var_ZLCD_HMI_bo_ZhangLi_CeDing_Adjustment")
      on Press: SetBit("ST_Var_ZLCD_HMI_bo_ZhangLi_CeDing_Adjustment")
   TextField "文本域_6" at 192,351 size 887x300; Text '张力弓整定步骤 1. 按下手动——>去使能 2. 拉住张力弓，同时按住停止和张力弓降两个按钮，卸去抱闸，将张力钢丝掉到走车撞块上 3. 按下手动按钮， 4. 点击张力测定，点击张力测定启动 5. 张力钢丝自动从最低点开始缓慢上升，同时自动记录数据 6. 待上升到48.5左右时张力弓停下 7. 观察以上6个数据，按下右侧的“调整”按钮，可看到前三个数据被第四个覆盖 8. 按下手动——>张力弓降，将张力钢丝降到正常位置 9. 结束'
   TextField "文本域_1" at 30,541 size 42x25; Text 'Text'

screen "保养提示" 1280x740, template "模板_根"
   on GenerateScreen: "TitleUpdater"()
   TextField "文本域_6" at 16,0 size 1000x680; Text '保养项目 已保养次数 1.锭子油更换:每隔 天,更换一次 2.龙带传动部分12个黄油嘴，加黄油（耐高温、高速、高负荷） 3.龙带压紧器，加黄油（耐高温 、高速、高负荷） 4.弓轴滚针轴承，每年加一次黄油 5.TC龙带，每两年清洗一次，水温小于15℃，阴凉通风处晾干 6.锭子传动同步带8M-2272 检查维护 7.控制柜清洁，三个月一次,用吸吹风机来吸内部粉尘 8.锭子电机风扇绕毛清理，两个月清理一次 9.其他，走车同步带轮、走车走轮绕毛定期检查清理'
   IOField "IO 域_3" at 836,87 size 65x39; FormatPattern 999
      ProcessValue <- "ST_Maintenance_g_u16_1_Times_OilChange_DingZi"
   IOField "IO 域_4" at 836,139 size 65x39; FormatPattern 999
      ProcessValue <- "ST_Maintenance_g_u16_2_Times_LongDai_HuangYouZui"
   IOField "IO 域_5" at 836,191 size 65x40; FormatPattern 999
      ProcessValue <- "ST_Maintenance_g_u16_3_Times_LongDai_YaJinQi"
   IOField "IO 域_6" at 836,244 size 65x39; FormatPattern 999
      ProcessValue <- "ST_Maintenance_g_u16_4_Times_GongZhou_Bearing"
   IOField "IO 域_7" at 836,296 size 65x39; FormatPattern 999
      ProcessValue <- "ST_Maintenance_g_u16_5_Times_LongDai_Clean"
   IOField "IO 域_8" at 836,348 size 65x40; FormatPattern 999
      ProcessValue <- "ST_Maintenance_g_u16_6_Times_DingZi_ChuanDong"
   IOField "IO 域_9" at 836,401 size 65x39; FormatPattern 999
      ProcessValue <- "ST_Maintenance_g_u16_7_Times_ControlBox_Clean"
   IOField "IO 域_10" at 836,453 size 65x39; FormatPattern 999
      ProcessValue <- "ST_Maintenance_g_u16_8_Times_DingZi_Fan"
   IOField "IO 域_1" at 258,87 size 66x39; Authorization "User administration"; FormatPattern 999
      ProcessValue <- "ST_Maintenance_g_u16_TimeInterval_OilChange"
   IOField "IO 域_2" at 486,15 size 65x39; Authorization "User administration"; FormatPattern 999
      ProcessValue <- "ST_Maintenance_g_u16_TimeReminder_Maintennance"
   TextField "文本域_4" at 317,19 size 160x35; Text '保养提醒持续'
   TextField "文本域_5" at 563,18 size 55x35; Text '天'
   Button "OBJECT_124" at 396,577 size 144x66; TextOn '罗拉关'; TextOff '罗拉开关 / EXIT'; Authorization "Operate_5"
      on Release: InvertBit("ST_Main_Var_ST_LuoLaSwitch")
      Appearance <- "ST_Main_Var_ST_LuoLaSwitch"

screen "报警管理" 1280x740, template "模板_根"
   on GenerateScreen: "TitleUpdater"()
   TextField "HmiScreenItemData_4" at 120,357 size 960x27; Text '报警画面'
   AlarmView "报警视图_1" at 0,0 size 1140x680; ColumnTextDevice 'D425 / PLC / API / ПЛК'; ColumnTextClassName '类别'; ColumnTextDiagnosable '可诊断'; ColumnTextNumber '编号 / No. / 番号 / 번호'
   Button "HmiScreenItemData_5" at 1150,396 size 130x47; TextOn '向后'; TextOff '报警记录'
      on Release: ActivateScreenByNumber("Picture", 0)
      on Press: SetTag("Picture", 61)
   Button "HmiScreenItemData_1" at 1150,314 size 130x47; TextOn '向后'; TextOff '监控画面'
      on Release: ActivateScreenByNumber("Picture", 0)
      on Press: SetTag("Picture", 62)

screen "报警记录" 1280x740, template "模板_根"
   on GenerateScreen: "TitleUpdater"()
   AlarmView "报警视图_1" at 0,0 size 1140x680; ColumnTextDevice 'D425 / PLC / API / ПЛК'
   Button "HmiScreenItemData_6" at 1150,396 size 130x47; TextOn '12张力弓整定'; TextOff '返回'
      on Release: ActivateScreenByNumber("Picture", 0); SetTag("ST_HMI_Var_HMI_i32_ZouChe_ZhanJu_ss_1", 0)
      on Press: SetTag("Picture", 6)

screen "车况设定" 1280x740, template "模板_设置"
   on GenerateScreen: "TitleUpdater"()
   TextField "Text Field_37" at 308,94 size 140x56; Text '出车展距:'
   TextField "Text Field_38" at 308,164 size 140x56; Text '出车速度:'
   TextField "Text Field_39" at 308,306 size 140x56; Text '进车速度:'
   TextField "Text Field_40" at 308,446 size 140x56; Text '出车时间:'
   TextField "Text Field_41" at 427,24 size 154x42; Text '车况设定'
   TextField "Text Field_42" at 308,516 size 140x56; Text '进车时间:'
   TextField "Text Field_43" at 672,94 size 84x56; Text 'mm'
   TextField "Text Field_44" at 672,164 size 84x56; Text 'mm/s'
   TextField "Text Field_45" at 672,306 size 84x56; Text 'mm/s'
   TextField "Text Field_46" at 672,446 size 84x56; Text '秒'
   TextField "Text Field_47" at 672,516 size 84x56; Text '秒'
   TextField "Text Field_48" at 266,234 size 182x56; Text '出车加速度:'
   TextField "Text Field_49" at 672,234 size 84x56; Text 'mm/s2'
   TextField "Text Field_50" at 252,376 size 196x56; Text '进车加速度:'
   TextField "Text Field_51" at 672,376 size 84x56; Text 'mm/s2'
   IOField "IO Field_20" at 504,94 size 140x56; FormatPattern 9999
      on OnFinishInput: SetBit("ST_Calculation_Var_HMI_bo_Calculation_0_Start")
      ProcessValue <- "ST_HMI_Var_HMI_r64Position_ChuChe"
   IOField "IO Field_21" at 504,164 size 140x56; FormatPattern 9999
      on OnFinishInput: SetBit("ST_Calculation_Var_HMI_bo_Calculation_0_Start")
      ProcessValue <- "ST_HMI_Var_HMI_r64Velocity_ChuChe"
   IOField "IO Field_22" at 504,306 size 140x56; FormatPattern 9999
      on OnFinishInput: SetBit("ST_Calculation_Var_HMI_bo_Calculation_0_Start")
      ProcessValue <- "ST_HMI_Var_HMI_r64Velocity_JinChe"
   IOField "IO Field_23" at 504,446 size 140x56; FormatPattern 99.9
      ProcessValue <- "ST_HMI_Var_HMI_r64Time_ChuChe"
      Appearance <- "ST_HMI_Var_HMI_boAlarm_NianDu_Time"
   IOField "IO Field_24" at 504,516 size 140x56; FormatPattern 99.9
      ProcessValue <- "ST_HMI_Var_HMI_r64Time_JinChe"
   IOField "IO Field_56" at 504,234 size 140x56; FormatPattern 9999
      ProcessValue <- "ST_HMI_Var_HMI_r64PositiveAccel_ZouChe_ChuChe"
   IOField "IO Field_70" at 504,376 size 140x56; FormatPattern 9999
      ProcessValue <- "ST_HMI_Var_HMI_r64PositiveAccel_ZouChe_JinChe"

screen "牵伸曲线" 1280x740, template "模板_设置"
   on GenerateScreen: "TitleUpdater"()
   TrendView "趋势视图_1" at 0,0 size 1050x680
      ValueAxis1End <- "ST_HMI_Var_HMI_r64Axis_ZouChe_Position_real"
      ValueAxis2End <- "ST_HMI_Var_HMI_r64QianShen_All_object"

screen "纱穗参数设定" 1280x740, template "模板_设置"
   on GenerateScreen: "TitleUpdater"()
   TextField "Text Field_50" at 206,234 size 187x56; Text '总高度:'
   TextField "Text Field_51" at 206,304 size 187x56; Text '上锥体高度:'
   TextField "Text Field_52" at 311,24 size 280x42; Text '纱穗参数设定'
   TextField "Text Field_53" at 206,374 size 187x56; Text '上锥体高度M:'
   TextField "Text Field_55" at 626,164 size 84x56; Text 'mm'
   TextField "Text Field_56" at 626,234 size 84x56; Text 'mm'
   TextField "Text Field_57" at 626,304 size 84x56; Text 'mm'
   TextField "Text Field_58" at 626,374 size 84x56; Text 'mm'
   TextField "Text Field_59" at 206,444 size 187x56; Text '最大直径:'
   TextField "Text Field_60" at 626,444 size 84x56; Text 'mm'
   TextField "Text Field_54" at 206,94 size 187x56; Text '起始点高度:'
   TextField "Text Field_61" at 626,94 size 84x56; Text 'mm'
   TextField "Text Field_62" at 206,164 size 187x56; Text '下锥体高度:'
   IOField "IO Field_27" at 444,234 size 140x56; FormatPattern 999.9
      ProcessValue <- "ST_HMI_Var_HMI_r64Height_ShaSui_whole"
   IOField "IO Field_28" at 444,304 size 140x56; FormatPattern 99.9
      ProcessValue <- "ST_HMI_Var_HMI_r64Height_ShaSui_Top"
   IOField "IO Field_29" at 444,374 size 140x56; FormatPattern 99.9
      ProcessValue <- "ST_HMI_Var_HMI_r64Height_ShaSui_Top_MaxD"
   IOField "IO Field_30" at 444,444 size 140x56; FormatPattern 99.9
      ProcessValue <- "ST_HMI_Var_HMI_r64Diameter_ShaSui_Max"
   IOField "IO Field_31" at 444,94 size 140x56; FormatPattern 99.9
      ProcessValue <- "ST_HMI_Var_HMI_r64Height_ShaSui_Start"
   IOField "IO Field_32" at 444,164 size 140x56; FormatPattern 99.9
      ProcessValue <- "ST_HMI_Var_HMI_r64Height_ShaSui_Bottom"
   TextField "Text Field_1" at 205,515 size 187x56; Text '纱管安装高度:'
   TextField "Text Field_2" at 625,515 size 84x56; Text 'mm'
   IOField "IO Field_1" at 443,515 size 140x56; FormatPattern 99.9
      ProcessValue <- "ST_HMI_Var_HMI_r64_h0_s"